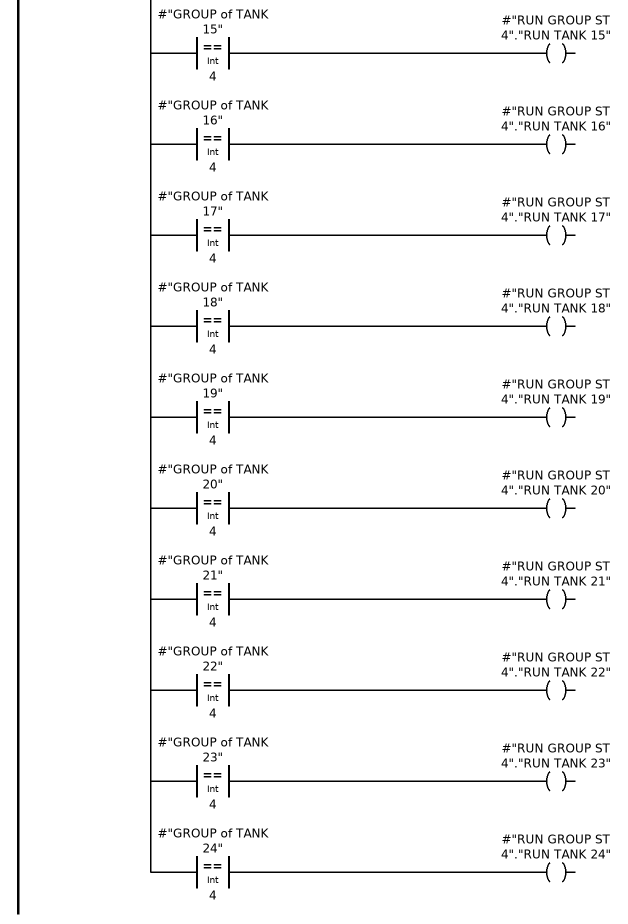
   RUNG wire#powerrail
      Contact( #"RUN GROUP 4" )
      wire#w1
      { S7_Templates := "SrcType := Int" } EQ_Contact(in1 := #"GROUP of TANK 1", in2 := 4)
      Coil( #"RUN GROUP ST 4"."RUN TANK 1" )
   END_RUNG
   RUNG wire#w1
      { S7_Templates := "SrcType := Int" } EQ_Contact(in1 := #"GROUP of TANK 2", in2 := 4)
      Coil( #"RUN GROUP ST 4"."RUN TANK 2" )
   END_RUNG
   RUNG wire#w1
      { S7_Templates := "SrcType := Int" } EQ_Contact(in1 := #"GROUP of TANK 3", in2 := 4)
      Coil( #"RUN GROUP ST 4"."RUN TANK 3" )
   END_RUNG
   RUNG wire#w1
      { S7_Templates := "SrcType := Int" } EQ_Contact(in1 := #"GROUP of TANK 4", in2 := 4)
      Coil( #"RUN GROUP ST 4"."RUN TANK 4" )
   END_RUNG
   RUNG wire#w1
      { S7_Templates := "SrcType := Int" } EQ_Contact(in1 := #"GROUP of TANK 5", in2 := 4)
      Coil( #"RUN GROUP ST 4"."RUN TANK 5" )
   END_RUNG
   RUNG wire#w1
      { S7_Templates := "SrcType := Int" } EQ_Contact(in1 := #"GROUP of TANK 6", in2 := 4)
      Coil( #"RUN GROUP ST 4"."RUN TANK 6" )
   END_RUNG
   RUNG wire#w1
      { S7_Templates := "SrcType := Int" } EQ_Contact(in1 := #"GROUP of TANK 7", in2 := 4)
      Coil( #"RUN GROUP ST 4"."RUN TANK 7" )
   END_RUNG
   RUNG wire#w1
      { S7_Templates := "SrcType := Int" } EQ_Contact(in1 := #"GROUP of TANK 8", in2 := 4)
      Coil( #"RUN GROUP ST 4"."RUN TANK 8" )
   END_RUNG
   RUNG wire#w1
      { S7_Templates := "SrcType := Int" } EQ_Contact(in1 := #"GROUP of TANK 9", in2 := 4)
      Coil( #"RUN GROUP ST 4"."RUN TANK 9" )
   END_RUNG
   RUNG wire#w1
      { S7_Templates := "SrcType := Int" } EQ_Contact(in1 := #"GROUP of TANK 10", in2 := 4)
      Coil( #"RUN GROUP ST 4"."RUN TANK 10" )
   END_RUNG
   RUNG wire#w1
      { S7_Templates := "SrcType := Int" } EQ_Contact(in1 := #"GROUP of TANK 11", in2 := 4)
      Coil( #"RUN GROUP ST 4"."RUN TANK 11" )
   END_RUNG
   RUNG wire#w1
      { S7_Templates := "SrcType := Int" } EQ_Contact(in1 := #"GROUP of TANK 12", in2 := 4)
      Coil( #"RUN GROUP ST 4"."RUN TANK 12" )
   END_RUNG
   RUNG wire#w1
      { S7_Templates := "SrcType := Int" } EQ_Contact(in1 := #"GROUP of TANK 13", in2 := 4)
      Coil( #"RUN GROUP ST 4"."RUN TANK 13" )
   END_RUNG
   RUNG wire#w1
      { S7_Templates := "SrcType := Int" } EQ_Contact(in1 := #"GROUP of TANK 14", in2 := 4)
      Coil( #"RUN GROUP ST 4"."RUN TANK 14" )
   END_RUNG
   RUNG wire#w1
      { S7_Templates := "SrcType := Int" } EQ_Contact(in1 := #"GROUP of TANK 15", in2 := 4)
      Coil( #"RUN GROUP ST 4"."RUN TANK 15" )
   END_RUNG
   RUNG wire#w1
      { S7_Templates := "SrcType := Int" } EQ_Contact(in1 := #"GROUP of TANK 16", in2 := 4)
      Coil( #"RUN GROUP ST 4"."RUN TANK 16" )
   END_RUNG
   RUNG wire#w1
      { S7_Templates := "SrcType := Int" } EQ_Contact(in1 := #"GROUP of TANK 17", in2 := 4)
      Coil( #"RUN GROUP ST 4"."RUN TANK 17" )
   END_RUNG
   RUNG wire#w1
      { S7_Templates := "SrcType := Int" } EQ_Contact(in1 := #"GROUP of TANK 18", in2 := 4)
      Coil( #"RUN GROUP ST 4"."RUN TANK 18" )
   END_RUNG
   RUNG wire#w1
      { S7_Templates := "SrcType := Int" } EQ_Contact(in1 := #"GROUP of TANK 19", in2 := 4)
      Coil( #"RUN GROUP ST 4"."RUN TANK 19" )
   END_RUNG
   RUNG wire#w1
      { S7_Templates := "SrcType := Int" } EQ_Contact(in1 := #"GROUP of TANK 20", in2 := 4)
      Coil( #"RUN GROUP ST 4"."RUN TANK 20" )
   END_RUNG
   RUNG wire#w1
      { S7_Templates := "SrcType := Int" } EQ_Contact(in1 := #"GROUP of TANK 21", in2 := 4)
      Coil( #"RUN GROUP ST 4"."RUN TANK 21" )
   END_RUNG
   RUNG wire#w1
      { S7_Templates := "SrcType := Int" } EQ_Contact(in1 := #"GROUP of TANK 22", in2 := 4)
      Coil( #"RUN GROUP ST 4"."RUN TANK 22" )
   END_RUNG
   RUNG wire#w1
      { S7_Templates := "SrcType := Int" } EQ_Contact(in1 := #"GROUP of TANK 23", in2 := 4)
      Coil( #"RUN GROUP ST 4"."RUN TANK 23" )
   END_RUNG
   RUNG wire#w1
      { S7_Templates := "SrcType := Int" } EQ_Contact(in1 := #"GROUP of TANK 24", in2 := 4)
      Coil( #"RUN GROUP ST 4"."RUN TANK 24" )
   END_RUNG
   // the same network as SCL:
   #"RUN GROUP ST 4"."RUN TANK 1" := #"RUN GROUP 4" AND (#"GROUP of TANK 1" = 4);
   #"RUN GROUP ST 4"."RUN TANK 2" := #"RUN GROUP 4" AND (#"GROUP of TANK 2" = 4);
   #"RUN GROUP ST 4"."RUN TANK 3" := #"RUN GROUP 4" AND (#"GROUP of TANK 3" = 4);
   #"RUN GROUP ST 4"."RUN TANK 4" := #"RUN GROUP 4" AND (#"GROUP of TANK 4" = 4);
   #"RUN GROUP ST 4"."RUN TANK 5" := #"RUN GROUP 4" AND (#"GROUP of TANK 5" = 4);
   #"RUN GROUP ST 4"."RUN TANK 6" := #"RUN GROUP 4" AND (#"GROUP of TANK 6" = 4);
   #"RUN GROUP ST 4"."RUN TANK 7" := #"RUN GROUP 4" AND (#"GROUP of TANK 7" = 4);
   #"RUN GROUP ST 4"."RUN TANK 8" := #"RUN GROUP 4" AND (#"GROUP of TANK 8" = 4);
   #"RUN GROUP ST 4"."RUN TANK 9" := #"RUN GROUP 4" AND (#"GROUP of TANK 9" = 4);
   #"RUN GROUP ST 4"."RUN TANK 10" := #"RUN GROUP 4" AND (#"GROUP of TANK 10" = 4);
   #"RUN GROUP ST 4"."RUN TANK 11" := #"RUN GROUP 4" AND (#"GROUP of TANK 11" = 4);
   #"RUN GROUP ST 4"."RUN TANK 12" := #"RUN GROUP 4" AND (#"GROUP of TANK 12" = 4);
   #"RUN GROUP ST 4"."RUN TANK 13" := #"RUN GROUP 4" AND (#"GROUP of TANK 13" = 4);
   #"RUN GROUP ST 4"."RUN TANK 14" := #"RUN GROUP 4" AND (#"GROUP of TANK 14" = 4);
   #"RUN GROUP ST 4"."RUN TANK 15" := #"RUN GROUP 4" AND (#"GROUP of TANK 15" = 4);
   #"RUN GROUP ST 4"."RUN TANK 16" := #"RUN GROUP 4" AND (#"GROUP of TANK 16" = 4);
   #"RUN GROUP ST 4"."RUN TANK 17" := #"RUN GROUP 4" AND (#"GROUP of TANK 17" = 4);
   #"RUN GROUP ST 4"."RUN TANK 18" := #"RUN GROUP 4" AND (#"GROUP of TANK 18" = 4);
   #"RUN GROUP ST 4"."RUN TANK 19" := #"RUN GROUP 4" AND (#"GROUP of TANK 19" = 4);
   #"RUN GROUP ST 4"."RUN TANK 20" := #"RUN GROUP 4" AND (#"GROUP of TANK 20" = 4);
   #"RUN GROUP ST 4"."RUN TANK 21" := #"RUN GROUP 4" AND (#"GROUP of TANK 21" = 4);
   #"RUN GROUP ST 4"."RUN TANK 22" := #"RUN GROUP 4" AND (#"GROUP of TANK 22" = 4);
   #"RUN GROUP ST 4"."RUN TANK 23" := #"RUN GROUP 4" AND (#"GROUP of TANK 23" = 4);
   #"RUN GROUP ST 4"."RUN TANK 24" := #"RUN GROUP 4" AND (#"GROUP of TANK 24" = 4);
END_REGION

REGION Network 53: RUN GROUP 5
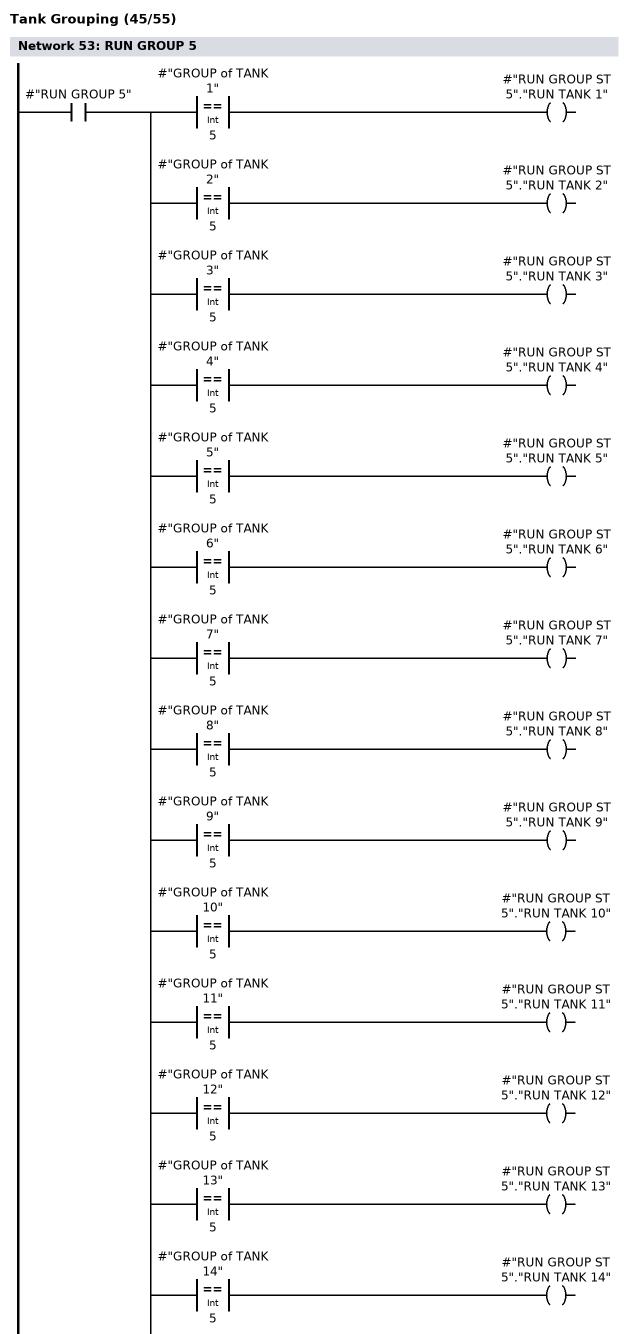
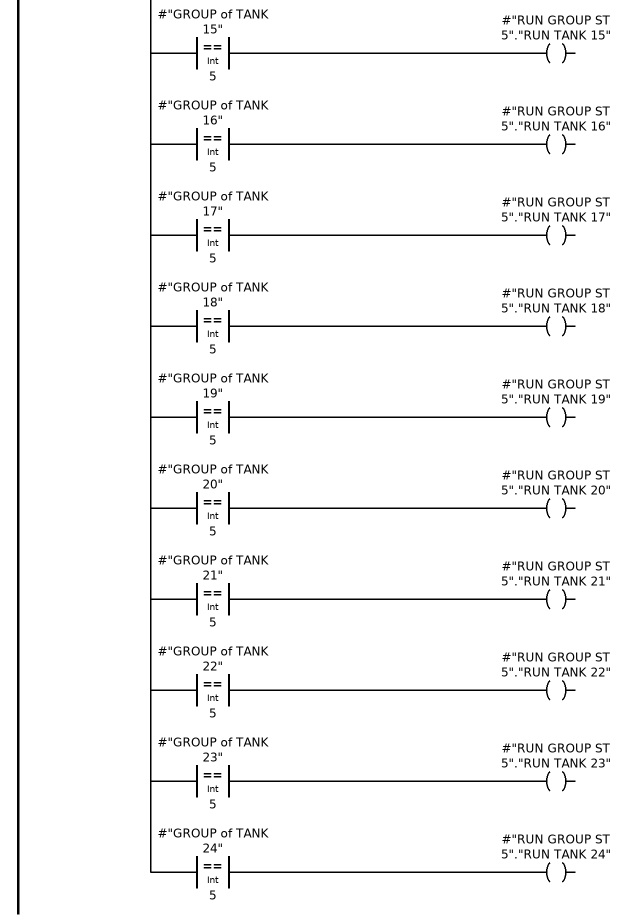
   RUNG wire#powerrail
      Contact( #"RUN GROUP 5" )
      wire#w1
      { S7_Templates := "SrcType := Int" } EQ_Contact(in1 := #"GROUP of TANK 1", in2 := 5)
      Coil( #"RUN GROUP ST 5"."RUN TANK 1" )
   END_RUNG
   RUNG wire#w1
      { S7_Templates := "SrcType := Int" } EQ_Contact(in1 := #"GROUP of TANK 2", in2 := 5)
      Coil( #"RUN GROUP ST 5"."RUN TANK 2" )
   END_RUNG
   RUNG wire#w1
      { S7_Templates := "SrcType := Int" } EQ_Contact(in1 := #"GROUP of TANK 3", in2 := 5)
      Coil( #"RUN GROUP ST 5"."RUN TANK 3" )
   END_RUNG
   RUNG wire#w1
      { S7_Templates := "SrcType := Int" } EQ_Contact(in1 := #"GROUP of TANK 4", in2 := 5)
      Coil( #"RUN GROUP ST 5"."RUN TANK 4" )
   END_RUNG
   RUNG wire#w1
      { S7_Templates := "SrcType := Int" } EQ_Contact(in1 := #"GROUP of TANK 5", in2 := 5)
      Coil( #"RUN GROUP ST 5"."RUN TANK 5" )
   END_RUNG
   RUNG wire#w1
      { S7_Templates := "SrcType := Int" } EQ_Contact(in1 := #"GROUP of TANK 6", in2 := 5)
      Coil( #"RUN GROUP ST 5"."RUN TANK 6" )
   END_RUNG
   RUNG wire#w1
      { S7_Templates := "SrcType := Int" } EQ_Contact(in1 := #"GROUP of TANK 7", in2 := 5)
      Coil( #"RUN GROUP ST 5"."RUN TANK 7" )
   END_RUNG
   RUNG wire#w1
      { S7_Templates := "SrcType := Int" } EQ_Contact(in1 := #"GROUP of TANK 8", in2 := 5)
      Coil( #"RUN GROUP ST 5"."RUN TANK 8" )
   END_RUNG
   RUNG wire#w1
      { S7_Templates := "SrcType := Int" } EQ_Contact(in1 := #"GROUP of TANK 9", in2 := 5)
      Coil( #"RUN GROUP ST 5"."RUN TANK 9" )
   END_RUNG
   RUNG wire#w1
      { S7_Templates := "SrcType := Int" } EQ_Contact(in1 := #"GROUP of TANK 10", in2 := 5)
      Coil( #"RUN GROUP ST 5"."RUN TANK 10" )
   END_RUNG
   RUNG wire#w1
      { S7_Templates := "SrcType := Int" } EQ_Contact(in1 := #"GROUP of TANK 11", in2 := 5)
      Coil( #"RUN GROUP ST 5"."RUN TANK 11" )
   END_RUNG
   RUNG wire#w1
      { S7_Templates := "SrcType := Int" } EQ_Contact(in1 := #"GROUP of TANK 12", in2 := 5)
      Coil( #"RUN GROUP ST 5"."RUN TANK 12" )
   END_RUNG
   RUNG wire#w1
      { S7_Templates := "SrcType := Int" } EQ_Contact(in1 := #"GROUP of TANK 13", in2 := 5)
      Coil( #"RUN GROUP ST 5"."RUN TANK 13" )
   END_RUNG
   RUNG wire#w1
      { S7_Templates := "SrcType := Int" } EQ_Contact(in1 := #"GROUP of TANK 14", in2 := 5)
      Coil( #"RUN GROUP ST 5"."RUN TANK 14" )
   END_RUNG
   RUNG wire#w1
      { S7_Templates := "SrcType := Int" } EQ_Contact(in1 := #"GROUP of TANK 15", in2 := 5)
      Coil( #"RUN GROUP ST 5"."RUN TANK 15" )
   END_RUNG
   RUNG wire#w1
      { S7_Templates := "SrcType := Int" } EQ_Contact(in1 := #"GROUP of TANK 16", in2 := 5)
      Coil( #"RUN GROUP ST 5"."RUN TANK 16" )
   END_RUNG
   RUNG wire#w1
      { S7_Templates := "SrcType := Int" } EQ_Contact(in1 := #"GROUP of TANK 17", in2 := 5)
      Coil( #"RUN GROUP ST 5"."RUN TANK 17" )
   END_RUNG
   RUNG wire#w1
      { S7_Templates := "SrcType := Int" } EQ_Contact(in1 := #"GROUP of TANK 18", in2 := 5)
      Coil( #"RUN GROUP ST 5"."RUN TANK 18" )
   END_RUNG
   RUNG wire#w1
      { S7_Templates := "SrcType := Int" } EQ_Contact(in1 := #"GROUP of TANK 19", in2 := 5)
      Coil( #"RUN GROUP ST 5"."RUN TANK 19" )
   END_RUNG
   RUNG wire#w1
      { S7_Templates := "SrcType := Int" } EQ_Contact(in1 := #"GROUP of TANK 20", in2 := 5)
      Coil( #"RUN GROUP ST 5"."RUN TANK 20" )
   END_RUNG
   RUNG wire#w1
      { S7_Templates := "SrcType := Int" } EQ_Contact(in1 := #"GROUP of TANK 21", in2 := 5)
      Coil( #"RUN GROUP ST 5"."RUN TANK 21" )
   END_RUNG
   RUNG wire#w1
      { S7_Templates := "SrcType := Int" } EQ_Contact(in1 := #"GROUP of TANK 22", in2 := 5)
      Coil( #"RUN GROUP ST 5"."RUN TANK 22" )
   END_RUNG
   RUNG wire#w1
      { S7_Templates := "SrcType := Int" } EQ_Contact(in1 := #"GROUP of TANK 23", in2 := 5)
      Coil( #"RUN GROUP ST 5"."RUN TANK 23" )
   END_RUNG
   RUNG wire#w1
      { S7_Templates := "SrcType := Int" } EQ_Contact(in1 := #"GROUP of TANK 24", in2 := 5)
      Coil( #"RUN GROUP ST 5"."RUN TANK 24" )
   END_RUNG
   // the same network as SCL:
   #"RUN GROUP ST 5"."RUN TANK 1" := #"RUN GROUP 5" AND (#"GROUP of TANK 1" = 5);
   #"RUN GROUP ST 5"."RUN TANK 2" := #"RUN GROUP 5" AND (#"GROUP of TANK 2" = 5);
   #"RUN GROUP ST 5"."RUN TANK 3" := #"RUN GROUP 5" AND (#"GROUP of TANK 3" = 5);
   #"RUN GROUP ST 5"."RUN TANK 4" := #"RUN GROUP 5" AND (#"GROUP of TANK 4" = 5);
   #"RUN GROUP ST 5"."RUN TANK 5" := #"RUN GROUP 5" AND (#"GROUP of TANK 5" = 5);
   #"RUN GROUP ST 5"."RUN TANK 6" := #"RUN GROUP 5" AND (#"GROUP of TANK 6" = 5);
   #"RUN GROUP ST 5"."RUN TANK 7" := #"RUN GROUP 5" AND (#"GROUP of TANK 7" = 5);
   #"RUN GROUP ST 5"."RUN TANK 8" := #"RUN GROUP 5" AND (#"GROUP of TANK 8" = 5);
   #"RUN GROUP ST 5"."RUN TANK 9" := #"RUN GROUP 5" AND (#"GROUP of TANK 9" = 5);
   #"RUN GROUP ST 5"."RUN TANK 10" := #"RUN GROUP 5" AND (#"GROUP of TANK 10" = 5);
   #"RUN GROUP ST 5"."RUN TANK 11" := #"RUN GROUP 5" AND (#"GROUP of TANK 11" = 5);
   #"RUN GROUP ST 5"."RUN TANK 12" := #"RUN GROUP 5" AND (#"GROUP of TANK 12" = 5);
   #"RUN GROUP ST 5"."RUN TANK 13" := #"RUN GROUP 5" AND (#"GROUP of TANK 13" = 5);
   #"RUN GROUP ST 5"."RUN TANK 14" := #"RUN GROUP 5" AND (#"GROUP of TANK 14" = 5);
   #"RUN GROUP ST 5"."RUN TANK 15" := #"RUN GROUP 5" AND (#"GROUP of TANK 15" = 5);
   #"RUN GROUP ST 5"."RUN TANK 16" := #"RUN GROUP 5" AND (#"GROUP of TANK 16" = 5);
   #"RUN GROUP ST 5"."RUN TANK 17" := #"RUN GROUP 5" AND (#"GROUP of TANK 17" = 5);
   #"RUN GROUP ST 5"."RUN TANK 18" := #"RUN GROUP 5" AND (#"GROUP of TANK 18" = 5);
   #"RUN GROUP ST 5"."RUN TANK 19" := #"RUN GROUP 5" AND (#"GROUP of TANK 19" = 5);
   #"RUN GROUP ST 5"."RUN TANK 20" := #"RUN GROUP 5" AND (#"GROUP of TANK 20" = 5);
   #"RUN GROUP ST 5"."RUN TANK 21" := #"RUN GROUP 5" AND (#"GROUP of TANK 21" = 5);
   #"RUN GROUP ST 5"."RUN TANK 22" := #"RUN GROUP 5" AND (#"GROUP of TANK 22" = 5);
   #"RUN GROUP ST 5"."RUN TANK 23" := #"RUN GROUP 5" AND (#"GROUP of TANK 23" = 5);
   #"RUN GROUP ST 5"."RUN TANK 24" := #"RUN GROUP 5" AND (#"GROUP of TANK 24" = 5);
END_REGION

REGION Network 54: RUN GROUP 6
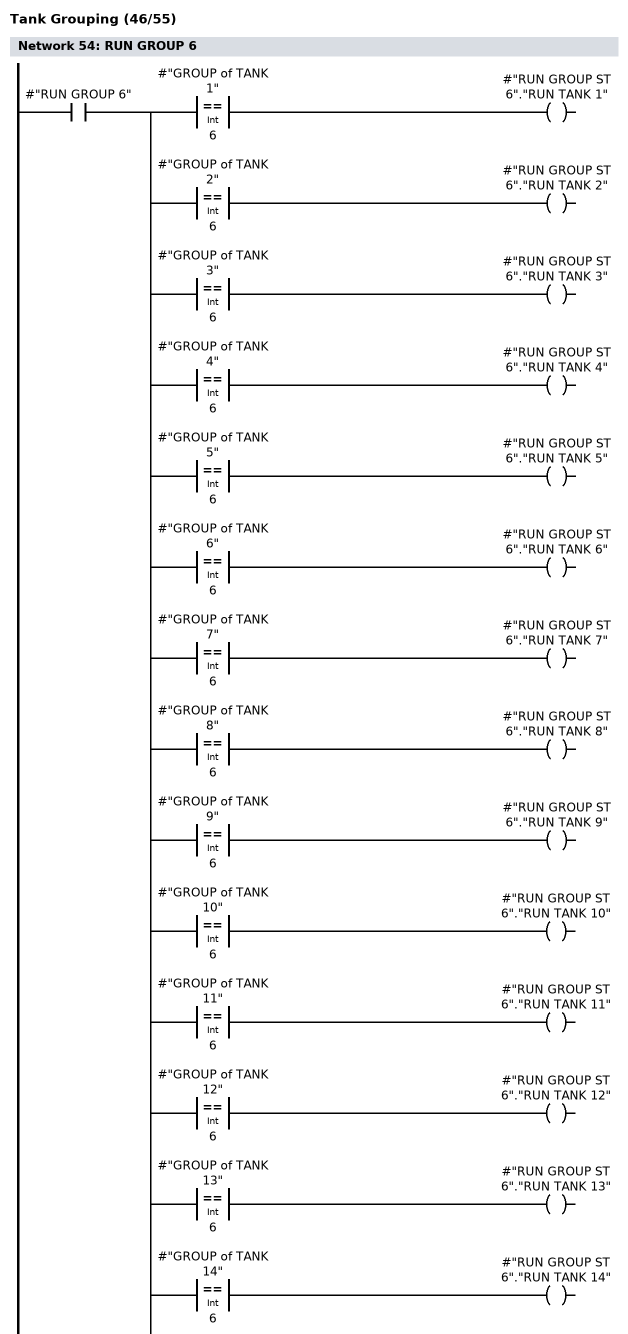
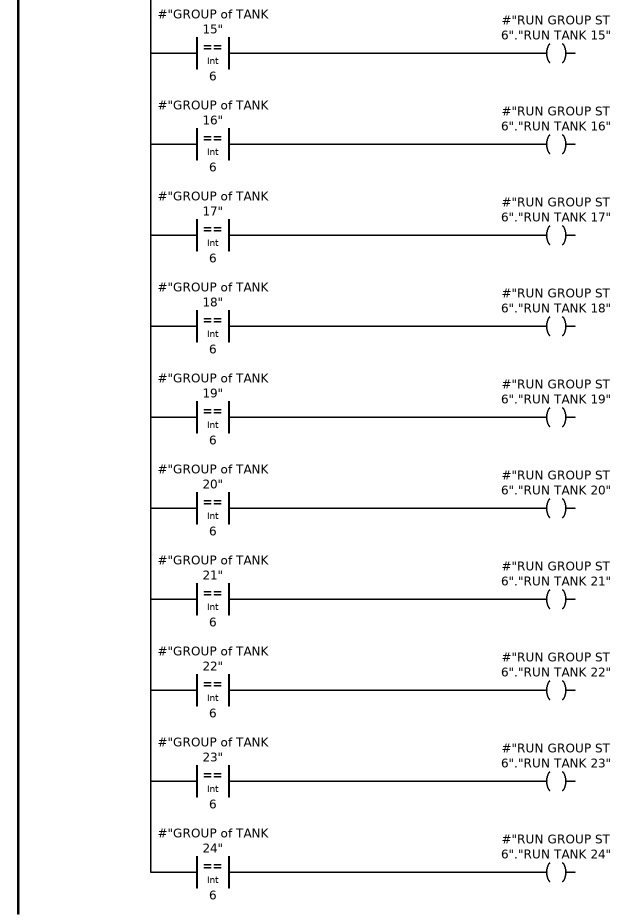
   RUNG wire#powerrail
      Contact( #"RUN GROUP 6" )
      wire#w1
      { S7_Templates := "SrcType := Int" } EQ_Contact(in1 := #"GROUP of TANK 1", in2 := 6)
      Coil( #"RUN GROUP ST 6"."RUN TANK 1" )
   END_RUNG
   RUNG wire#w1
      { S7_Templates := "SrcType := Int" } EQ_Contact(in1 := #"GROUP of TANK 2", in2 := 6)
      Coil( #"RUN GROUP ST 6"."RUN TANK 2" )
   END_RUNG
   RUNG wire#w1
      { S7_Templates := "SrcType := Int" } EQ_Contact(in1 := #"GROUP of TANK 3", in2 := 6)
      Coil( #"RUN GROUP ST 6"."RUN TANK 3" )
   END_RUNG
   RUNG wire#w1
      { S7_Templates := "SrcType := Int" } EQ_Contact(in1 := #"GROUP of TANK 4", in2 := 6)
      Coil( #"RUN GROUP ST 6"."RUN TANK 4" )
   END_RUNG
   RUNG wire#w1
      { S7_Templates := "SrcType := Int" } EQ_Contact(in1 := #"GROUP of TANK 5", in2 := 6)
      Coil( #"RUN GROUP ST 6"."RUN TANK 5" )
   END_RUNG
   RUNG wire#w1
      { S7_Templates := "SrcType := Int" } EQ_Contact(in1 := #"GROUP of TANK 6", in2 := 6)
      Coil( #"RUN GROUP ST 6"."RUN TANK 6" )
   END_RUNG
   RUNG wire#w1
      { S7_Templates := "SrcType := Int" } EQ_Contact(in1 := #"GROUP of TANK 7", in2 := 6)
      Coil( #"RUN GROUP ST 6"."RUN TANK 7" )
   END_RUNG
   RUNG wire#w1
      { S7_Templates := "SrcType := Int" } EQ_Contact(in1 := #"GROUP of TANK 8", in2 := 6)
      Coil( #"RUN GROUP ST 6"."RUN TANK 8" )
   END_RUNG
   RUNG wire#w1
      { S7_Templates := "SrcType := Int" } EQ_Contact(in1 := #"GROUP of TANK 9", in2 := 6)
      Coil( #"RUN GROUP ST 6"."RUN TANK 9" )
   END_RUNG
   RUNG wire#w1
      { S7_Templates := "SrcType := Int" } EQ_Contact(in1 := #"GROUP of TANK 10", in2 := 6)
      Coil( #"RUN GROUP ST 6"."RUN TANK 10" )
   END_RUNG
   RUNG wire#w1
      { S7_Templates := "SrcType := Int" } EQ_Contact(in1 := #"GROUP of TANK 11", in2 := 6)
      Coil( #"RUN GROUP ST 6"."RUN TANK 11" )
   END_RUNG
   RUNG wire#w1
      { S7_Templates := "SrcType := Int" } EQ_Contact(in1 := #"GROUP of TANK 12", in2 := 6)
      Coil( #"RUN GROUP ST 6"."RUN TANK 12" )
   END_RUNG
   RUNG wire#w1
      { S7_Templates := "SrcType := Int" } EQ_Contact(in1 := #"GROUP of TANK 13", in2 := 6)
      Coil( #"RUN GROUP ST 6"."RUN TANK 13" )
   END_RUNG
   RUNG wire#w1
      { S7_Templates := "SrcType := Int" } EQ_Contact(in1 := #"GROUP of TANK 14", in2 := 6)
      Coil( #"RUN GROUP ST 6"."RUN TANK 14" )
   END_RUNG
   RUNG wire#w1
      { S7_Templates := "SrcType := Int" } EQ_Contact(in1 := #"GROUP of TANK 15", in2 := 6)
      Coil( #"RUN GROUP ST 6"."RUN TANK 15" )
   END_RUNG
   RUNG wire#w1
      { S7_Templates := "SrcType := Int" } EQ_Contact(in1 := #"GROUP of TANK 16", in2 := 6)
      Coil( #"RUN GROUP ST 6"."RUN TANK 16" )
   END_RUNG
   RUNG wire#w1
      { S7_Templates := "SrcType := Int" } EQ_Contact(in1 := #"GROUP of TANK 17", in2 := 6)
      Coil( #"RUN GROUP ST 6"."RUN TANK 17" )
   END_RUNG
   RUNG wire#w1
      { S7_Templates := "SrcType := Int" } EQ_Contact(in1 := #"GROUP of TANK 18", in2 := 6)
      Coil( #"RUN GROUP ST 6"."RUN TANK 18" )
   END_RUNG
   RUNG wire#w1
      { S7_Templates := "SrcType := Int" } EQ_Contact(in1 := #"GROUP of TANK 19", in2 := 6)
      Coil( #"RUN GROUP ST 6"."RUN TANK 19" )
   END_RUNG
   RUNG wire#w1
      { S7_Templates := "SrcType := Int" } EQ_Contact(in1 := #"GROUP of TANK 20", in2 := 6)
      Coil( #"RUN GROUP ST 6"."RUN TANK 20" )
   END_RUNG
   RUNG wire#w1
      { S7_Templates := "SrcType := Int" } EQ_Contact(in1 := #"GROUP of TANK 21", in2 := 6)
      Coil( #"RUN GROUP ST 6"."RUN TANK 21" )
   END_RUNG
   RUNG wire#w1
      { S7_Templates := "SrcType := Int" } EQ_Contact(in1 := #"GROUP of TANK 22", in2 := 6)
      Coil( #"RUN GROUP ST 6"."RUN TANK 22" )
   END_RUNG
   RUNG wire#w1
      { S7_Templates := "SrcType := Int" } EQ_Contact(in1 := #"GROUP of TANK 23", in2 := 6)
      Coil( #"RUN GROUP ST 6"."RUN TANK 23" )
   END_RUNG
   RUNG wire#w1
      { S7_Templates := "SrcType := Int" } EQ_Contact(in1 := #"GROUP of TANK 24", in2 := 6)
      Coil( #"RUN GROUP ST 6"."RUN TANK 24" )
   END_RUNG
   // the same network as SCL:
   #"RUN GROUP ST 6"."RUN TANK 1" := #"RUN GROUP 6" AND (#"GROUP of TANK 1" = 6);
   #"RUN GROUP ST 6"."RUN TANK 2" := #"RUN GROUP 6" AND (#"GROUP of TANK 2" = 6);
   #"RUN GROUP ST 6"."RUN TANK 3" := #"RUN GROUP 6" AND (#"GROUP of TANK 3" = 6);
   #"RUN GROUP ST 6"."RUN TANK 4" := #"RUN GROUP 6" AND (#"GROUP of TANK 4" = 6);
   #"RUN GROUP ST 6"."RUN TANK 5" := #"RUN GROUP 6" AND (#"GROUP of TANK 5" = 6);
   #"RUN GROUP ST 6"."RUN TANK 6" := #"RUN GROUP 6" AND (#"GROUP of TANK 6" = 6);
   #"RUN GROUP ST 6"."RUN TANK 7" := #"RUN GROUP 6" AND (#"GROUP of TANK 7" = 6);
   #"RUN GROUP ST 6"."RUN TANK 8" := #"RUN GROUP 6" AND (#"GROUP of TANK 8" = 6);
   #"RUN GROUP ST 6"."RUN TANK 9" := #"RUN GROUP 6" AND (#"GROUP of TANK 9" = 6);
   #"RUN GROUP ST 6"."RUN TANK 10" := #"RUN GROUP 6" AND (#"GROUP of TANK 10" = 6);
   #"RUN GROUP ST 6"."RUN TANK 11" := #"RUN GROUP 6" AND (#"GROUP of TANK 11" = 6);
   #"RUN GROUP ST 6"."RUN TANK 12" := #"RUN GROUP 6" AND (#"GROUP of TANK 12" = 6);
   #"RUN GROUP ST 6"."RUN TANK 13" := #"RUN GROUP 6" AND (#"GROUP of TANK 13" = 6);
   #"RUN GROUP ST 6"."RUN TANK 14" := #"RUN GROUP 6" AND (#"GROUP of TANK 14" = 6);
   #"RUN GROUP ST 6"."RUN TANK 15" := #"RUN GROUP 6" AND (#"GROUP of TANK 15" = 6);
   #"RUN GROUP ST 6"."RUN TANK 16" := #"RUN GROUP 6" AND (#"GROUP of TANK 16" = 6);
   #"RUN GROUP ST 6"."RUN TANK 17" := #"RUN GROUP 6" AND (#"GROUP of TANK 17" = 6);
   #"RUN GROUP ST 6"."RUN TANK 18" := #"RUN GROUP 6" AND (#"GROUP of TANK 18" = 6);
   #"RUN GROUP ST 6"."RUN TANK 19" := #"RUN GROUP 6" AND (#"GROUP of TANK 19" = 6);
   #"RUN GROUP ST 6"."RUN TANK 20" := #"RUN GROUP 6" AND (#"GROUP of TANK 20" = 6);
   #"RUN GROUP ST 6"."RUN TANK 21" := #"RUN GROUP 6" AND (#"GROUP of TANK 21" = 6);
   #"RUN GROUP ST 6"."RUN TANK 22" := #"RUN GROUP 6" AND (#"GROUP of TANK 22" = 6);
   #"RUN GROUP ST 6"."RUN TANK 23" := #"RUN GROUP 6" AND (#"GROUP of TANK 23" = 6);
   #"RUN GROUP ST 6"."RUN TANK 24" := #"RUN GROUP 6" AND (#"GROUP of TANK 24" = 6);
END_REGION

REGION Network 55: RUN GROUP 7
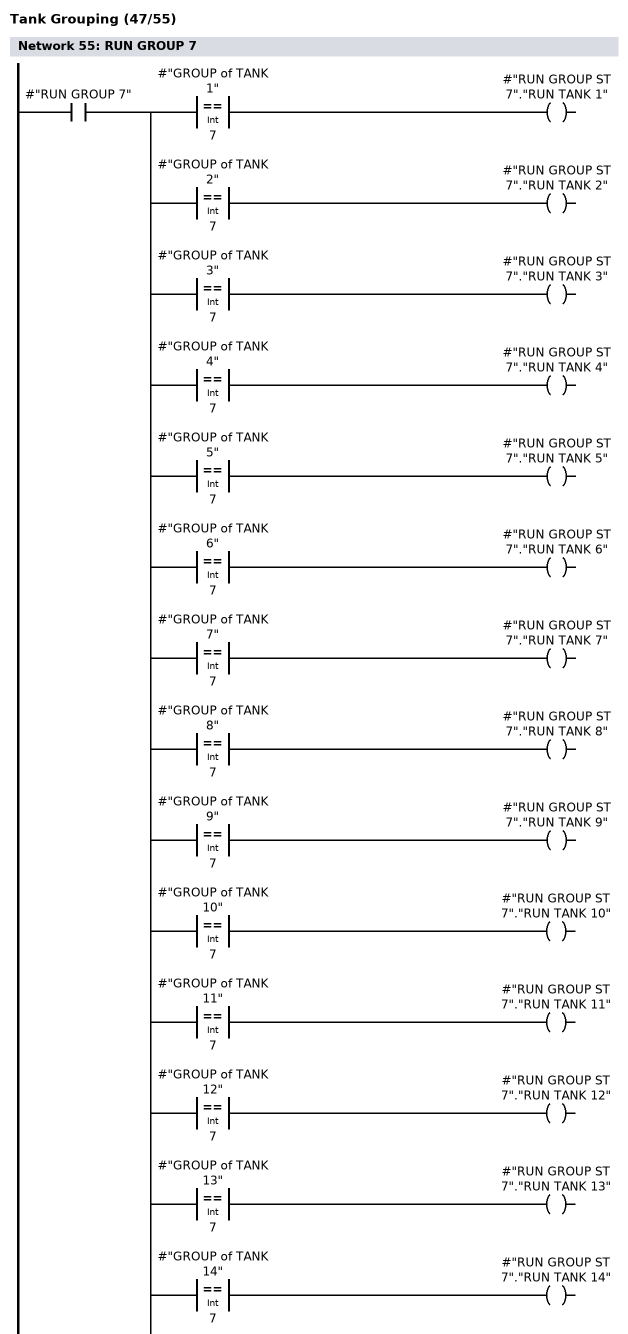
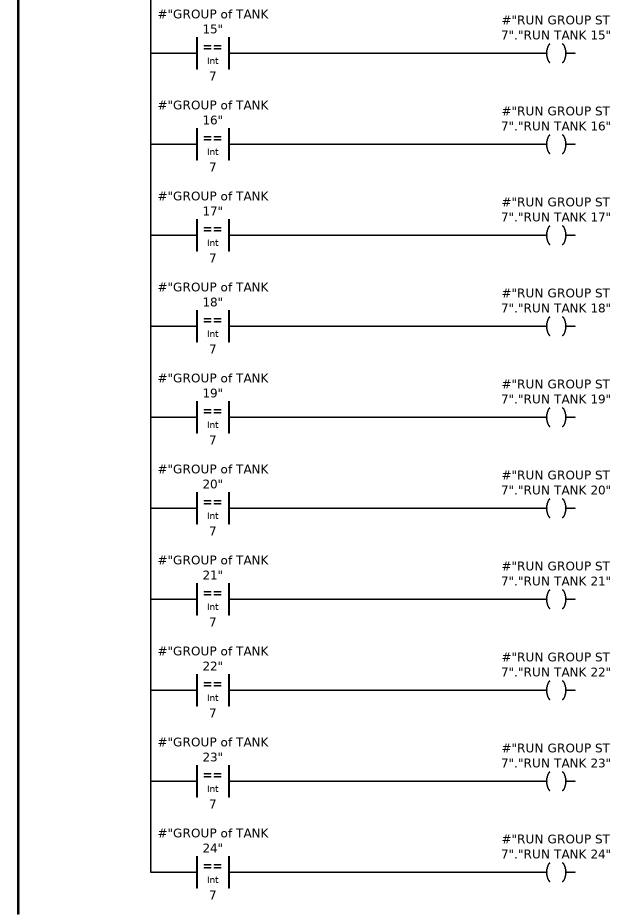
   RUNG wire#powerrail
      Contact( #"RUN GROUP 7" )
      wire#w1
      { S7_Templates := "SrcType := Int" } EQ_Contact(in1 := #"GROUP of TANK 1", in2 := 7)
      Coil( #"RUN GROUP ST 7"."RUN TANK 1" )
   END_RUNG
   RUNG wire#w1
      { S7_Templates := "SrcType := Int" } EQ_Contact(in1 := #"GROUP of TANK 2", in2 := 7)
      Coil( #"RUN GROUP ST 7"."RUN TANK 2" )
   END_RUNG
   RUNG wire#w1
      { S7_Templates := "SrcType := Int" } EQ_Contact(in1 := #"GROUP of TANK 3", in2 := 7)
      Coil( #"RUN GROUP ST 7"."RUN TANK 3" )
   END_RUNG
   RUNG wire#w1
      { S7_Templates := "SrcType := Int" } EQ_Contact(in1 := #"GROUP of TANK 4", in2 := 7)
      Coil( #"RUN GROUP ST 7"."RUN TANK 4" )
   END_RUNG
   RUNG wire#w1
      { S7_Templates := "SrcType := Int" } EQ_Contact(in1 := #"GROUP of TANK 5", in2 := 7)
      Coil( #"RUN GROUP ST 7"."RUN TANK 5" )
   END_RUNG
   RUNG wire#w1
      { S7_Templates := "SrcType := Int" } EQ_Contact(in1 := #"GROUP of TANK 6", in2 := 7)
      Coil( #"RUN GROUP ST 7"."RUN TANK 6" )
   END_RUNG
   RUNG wire#w1
      { S7_Templates := "SrcType := Int" } EQ_Contact(in1 := #"GROUP of TANK 7", in2 := 7)
      Coil( #"RUN GROUP ST 7"."RUN TANK 7" )
   END_RUNG
   RUNG wire#w1
      { S7_Templates := "SrcType := Int" } EQ_Contact(in1 := #"GROUP of TANK 8", in2 := 7)
      Coil( #"RUN GROUP ST 7"."RUN TANK 8" )
   END_RUNG
   RUNG wire#w1
      { S7_Templates := "SrcType := Int" } EQ_Contact(in1 := #"GROUP of TANK 9", in2 := 7)
      Coil( #"RUN GROUP ST 7"."RUN TANK 9" )
   END_RUNG
   RUNG wire#w1
      { S7_Templates := "SrcType := Int" } EQ_Contact(in1 := #"GROUP of TANK 10", in2 := 7)
      Coil( #"RUN GROUP ST 7"."RUN TANK 10" )
   END_RUNG
   RUNG wire#w1
      { S7_Templates := "SrcType := Int" } EQ_Contact(in1 := #"GROUP of TANK 11", in2 := 7)
      Coil( #"RUN GROUP ST 7"."RUN TANK 11" )
   END_RUNG
   RUNG wire#w1
      { S7_Templates := "SrcType := Int" } EQ_Contact(in1 := #"GROUP of TANK 12", in2 := 7)
      Coil( #"RUN GROUP ST 7"."RUN TANK 12" )
   END_RUNG
   RUNG wire#w1
      { S7_Templates := "SrcType := Int" } EQ_Contact(in1 := #"GROUP of TANK 13", in2 := 7)
      Coil( #"RUN GROUP ST 7"."RUN TANK 13" )
   END_RUNG
   RUNG wire#w1
      { S7_Templates := "SrcType := Int" } EQ_Contact(in1 := #"GROUP of TANK 14", in2 := 7)
      Coil( #"RUN GROUP ST 7"."RUN TANK 14" )
   END_RUNG
   RUNG wire#w1
      { S7_Templates := "SrcType := Int" } EQ_Contact(in1 := #"GROUP of TANK 15", in2 := 7)
      Coil( #"RUN GROUP ST 7"."RUN TANK 15" )
   END_RUNG
   RUNG wire#w1
      { S7_Templates := "SrcType := Int" } EQ_Contact(in1 := #"GROUP of TANK 16", in2 := 7)
      Coil( #"RUN GROUP ST 7"."RUN TANK 16" )
   END_RUNG
   RUNG wire#w1
      { S7_Templates := "SrcType := Int" } EQ_Contact(in1 := #"GROUP of TANK 17", in2 := 7)
      Coil( #"RUN GROUP ST 7"."RUN TANK 17" )
   END_RUNG
   RUNG wire#w1
      { S7_Templates := "SrcType := Int" } EQ_Contact(in1 := #"GROUP of TANK 18", in2 := 7)
      Coil( #"RUN GROUP ST 7"."RUN TANK 18" )
   END_RUNG
   RUNG wire#w1
      { S7_Templates := "SrcType := Int" } EQ_Contact(in1 := #"GROUP of TANK 19", in2 := 7)
      Coil( #"RUN GROUP ST 7"."RUN TANK 19" )
   END_RUNG
   RUNG wire#w1
      { S7_Templates := "SrcType := Int" } EQ_Contact(in1 := #"GROUP of TANK 20", in2 := 7)
      Coil( #"RUN GROUP ST 7"."RUN TANK 20" )
   END_RUNG
   RUNG wire#w1
      { S7_Templates := "SrcType := Int" } EQ_Contact(in1 := #"GROUP of TANK 21", in2 := 7)
      Coil( #"RUN GROUP ST 7"."RUN TANK 21" )
   END_RUNG
   RUNG wire#w1
      { S7_Templates := "SrcType := Int" } EQ_Contact(in1 := #"GROUP of TANK 22", in2 := 7)
      Coil( #"RUN GROUP ST 7"."RUN TANK 22" )
   END_RUNG
   RUNG wire#w1
      { S7_Templates := "SrcType := Int" } EQ_Contact(in1 := #"GROUP of TANK 23", in2 := 7)
      Coil( #"RUN GROUP ST 7"."RUN TANK 23" )
   END_RUNG
   RUNG wire#w1
      { S7_Templates := "SrcType := Int" } EQ_Contact(in1 := #"GROUP of TANK 24", in2 := 7)
      Coil( #"RUN GROUP ST 7"."RUN TANK 24" )
   END_RUNG
   // the same network as SCL:
   #"RUN GROUP ST 7"."RUN TANK 1" := #"RUN GROUP 7" AND (#"GROUP of TANK 1" = 7);
   #"RUN GROUP ST 7"."RUN TANK 2" := #"RUN GROUP 7" AND (#"GROUP of TANK 2" = 7);
   #"RUN GROUP ST 7"."RUN TANK 3" := #"RUN GROUP 7" AND (#"GROUP of TANK 3" = 7);
   #"RUN GROUP ST 7"."RUN TANK 4" := #"RUN GROUP 7" AND (#"GROUP of TANK 4" = 7);
   #"RUN GROUP ST 7"."RUN TANK 5" := #"RUN GROUP 7" AND (#"GROUP of TANK 5" = 7);
   #"RUN GROUP ST 7"."RUN TANK 6" := #"RUN GROUP 7" AND (#"GROUP of TANK 6" = 7);
   #"RUN GROUP ST 7"."RUN TANK 7" := #"RUN GROUP 7" AND (#"GROUP of TANK 7" = 7);
   #"RUN GROUP ST 7"."RUN TANK 8" := #"RUN GROUP 7" AND (#"GROUP of TANK 8" = 7);
   #"RUN GROUP ST 7"."RUN TANK 9" := #"RUN GROUP 7" AND (#"GROUP of TANK 9" = 7);
   #"RUN GROUP ST 7"."RUN TANK 10" := #"RUN GROUP 7" AND (#"GROUP of TANK 10" = 7);
   #"RUN GROUP ST 7"."RUN TANK 11" := #"RUN GROUP 7" AND (#"GROUP of TANK 11" = 7);
   #"RUN GROUP ST 7"."RUN TANK 12" := #"RUN GROUP 7" AND (#"GROUP of TANK 12" = 7);
   #"RUN GROUP ST 7"."RUN TANK 13" := #"RUN GROUP 7" AND (#"GROUP of TANK 13" = 7);
   #"RUN GROUP ST 7"."RUN TANK 14" := #"RUN GROUP 7" AND (#"GROUP of TANK 14" = 7);
   #"RUN GROUP ST 7"."RUN TANK 15" := #"RUN GROUP 7" AND (#"GROUP of TANK 15" = 7);
   #"RUN GROUP ST 7"."RUN TANK 16" := #"RUN GROUP 7" AND (#"GROUP of TANK 16" = 7);
   #"RUN GROUP ST 7"."RUN TANK 17" := #"RUN GROUP 7" AND (#"GROUP of TANK 17" = 7);
   #"RUN GROUP ST 7"."RUN TANK 18" := #"RUN GROUP 7" AND (#"GROUP of TANK 18" = 7);
   #"RUN GROUP ST 7"."RUN TANK 19" := #"RUN GROUP 7" AND (#"GROUP of TANK 19" = 7);
   #"RUN GROUP ST 7"."RUN TANK 20" := #"RUN GROUP 7" AND (#"GROUP of TANK 20" = 7);
   #"RUN GROUP ST 7"."RUN TANK 21" := #"RUN GROUP 7" AND (#"GROUP of TANK 21" = 7);
   #"RUN GROUP ST 7"."RUN TANK 22" := #"RUN GROUP 7" AND (#"GROUP of TANK 22" = 7);
   #"RUN GROUP ST 7"."RUN TANK 23" := #"RUN GROUP 7" AND (#"GROUP of TANK 23" = 7);
   #"RUN GROUP ST 7"."RUN TANK 24" := #"RUN GROUP 7" AND (#"GROUP of TANK 24" = 7);
END_REGION

REGION Network 56: RUN GROUP 8